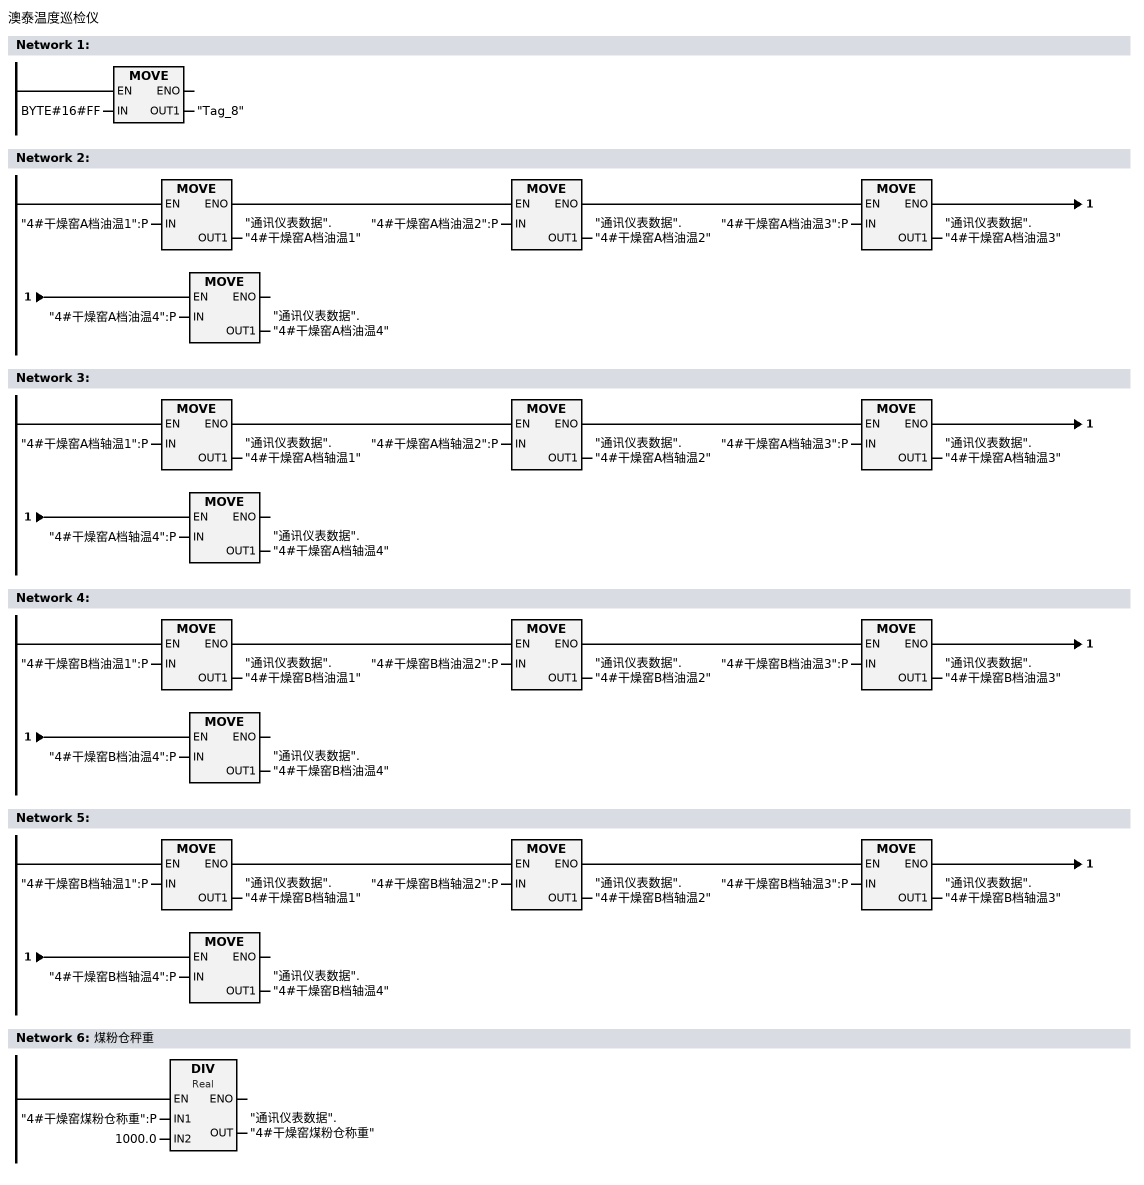
   RUNG wire#powerrail
      { S7_GenerateENO := "TRUE" } Move(in := BYTE#16#FF, out1 => "Tag_8")
   END_RUNG
   // the same network as SCL:
   "Tag_8" := BYTE#16#FF;
END_REGION

REGION Network 2
   RUNG wire#powerrail
      { S7_GenerateENO := "TRUE" } Move(in := "4#干燥窑A档油温1":P, out1 => "通讯仪表数据"."4#干燥窑A档油温1")
      { S7_GenerateENO := "TRUE" } Move(in := "4#干燥窑A档油温2":P, out1 => "通讯仪表数据"."4#干燥窑A档油温2")
      { S7_GenerateENO := "TRUE" } Move(in := "4#干燥窑A档油温3":P, out1 => "通讯仪表数据"."4#干燥窑A档油温3")
      { S7_GenerateENO := "TRUE" } Move(in := "4#干燥窑A档油温4":P, out1 => "通讯仪表数据"."4#干燥窑A档油温4")
   END_RUNG
   // the same network as SCL:
   // ENO of a box is taken as its EN; it also drops when the box reports an error
   "通讯仪表数据"."4#干燥窑A档油温1" := "4#干燥窑A档油温1":P;
   "通讯仪表数据"."4#干燥窑A档油温2" := "4#干燥窑A档油温2":P;
   "通讯仪表数据"."4#干燥窑A档油温3" := "4#干燥窑A档油温3":P;
   "通讯仪表数据"."4#干燥窑A档油温4" := "4#干燥窑A档油温4":P;
END_REGION

REGION Network 3
   RUNG wire#powerrail
      { S7_GenerateENO := "TRUE" } Move(in := "4#干燥窑A档轴温1":P, out1 => "通讯仪表数据"."4#干燥窑A档轴温1")
      { S7_GenerateENO := "TRUE" } Move(in := "4#干燥窑A档轴温2":P, out1 => "通讯仪表数据"."4#干燥窑A档轴温2")
      { S7_GenerateENO := "TRUE" } Move(in := "4#干燥窑A档轴温3":P, out1 => "通讯仪表数据"."4#干燥窑A档轴温3")
      { S7_GenerateENO := "TRUE" } Move(in := "4#干燥窑A档轴温4":P, out1 => "通讯仪表数据"."4#干燥窑A档轴温4")
   END_RUNG
   // the same network as SCL:
   // ENO of a box is taken as its EN; it also drops when the box reports an error
   "通讯仪表数据"."4#干燥窑A档轴温1" := "4#干燥窑A档轴温1":P;
   "通讯仪表数据"."4#干燥窑A档轴温2" := "4#干燥窑A档轴温2":P;
   "通讯仪表数据"."4#干燥窑A档轴温3" := "4#干燥窑A档轴温3":P;
   "通讯仪表数据"."4#干燥窑A档轴温4" := "4#干燥窑A档轴温4":P;
END_REGION

REGION Network 4
   RUNG wire#powerrail
      { S7_GenerateENO := "TRUE" } Move(in := "4#干燥窑B档油温1":P, out1 => "通讯仪表数据"."4#干燥窑B档油温1")
      { S7_GenerateENO := "TRUE" } Move(in := "4#干燥窑B档油温2":P, out1 => "通讯仪表数据"."4#干燥窑B档油温2")
      { S7_GenerateENO := "TRUE" } Move(in := "4#干燥窑B档油温3":P, out1 => "通讯仪表数据"."4#干燥窑B档油温3")
      { S7_GenerateENO := "TRUE" } Move(in := "4#干燥窑B档油温4":P, out1 => "通讯仪表数据"."4#干燥窑B档油温4")
   END_RUNG
   // the same network as SCL:
   // ENO of a box is taken as its EN; it also drops when the box reports an error
   "通讯仪表数据"."4#干燥窑B档油温1" := "4#干燥窑B档油温1":P;
   "通讯仪表数据"."4#干燥窑B档油温2" := "4#干燥窑B档油温2":P;
   "通讯仪表数据"."4#干燥窑B档油温3" := "4#干燥窑B档油温3":P;
   "通讯仪表数据"."4#干燥窑B档油温4" := "4#干燥窑B档油温4":P;
END_REGION

REGION Network 5
   RUNG wire#powerrail
      { S7_GenerateENO := "TRUE" } Move(in := "4#干燥窑B档轴温1":P, out1 => "通讯仪表数据"."4#干燥窑B档轴温1")
      { S7_GenerateENO := "TRUE" } Move(in := "4#干燥窑B档轴温2":P, out1 => "通讯仪表数据"."4#干燥窑B档轴温2")
      { S7_GenerateENO := "TRUE" } Move(in := "4#干燥窑B档轴温3":P, out1 => "通讯仪表数据"."4#干燥窑B档轴温3")
      { S7_GenerateENO := "TRUE" } Move(in := "4#干燥窑B档轴温4":P, out1 => "通讯仪表数据"."4#干燥窑B档轴温4")
   END_RUNG
   // the same network as SCL:
   // ENO of a box is taken as its EN; it also drops when the box reports an error
   "通讯仪表数据"."4#干燥窑B档轴温1" := "4#干燥窑B档轴温1":P;
   "通讯仪表数据"."4#干燥窑B档轴温2" := "4#干燥窑B档轴温2":P;
   "通讯仪表数据"."4#干燥窑B档轴温3" := "4#干燥窑B档轴温3":P;
   "通讯仪表数据"."4#干燥窑B档轴温4" := "4#干燥窑B档轴温4":P;
END_REGION

REGION Network 6: 煤粉仓秤重
   RUNG wire#powerrail
      { S7_Templates := "SrcType := Real" } Div(in1 := "4#干燥窑煤粉仓称重":P, in2 := 1000.0, out => "通讯仪表数据"."4#干燥窑煤粉仓称重")
   END_RUNG
   // the same network as SCL:
   "通讯仪表数据"."4#干燥窑煤粉仓称重" := "4#干燥窑煤粉仓称重":P / 1000.0;
END_REGION
END_FUNCTION

FUNCTION "3#4#干燥窑皮带联锁信号通" : Void   // FC16, LAD
{ S7_Optimized_Access := 'FALSE' }
VERSION : 0.1
BEGIN

REGION Network 1
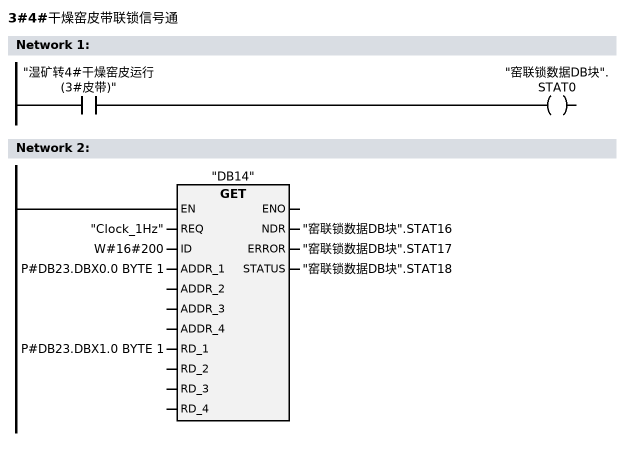
   RUNG wire#powerrail
      Contact( "湿矿转4#干燥窑皮运行  (3#皮带)" )
      Coil( "窑联锁数据DB块".STAT0 )
   END_RUNG
   // the same network as SCL:
   "窑联锁数据DB块".STAT0 := "湿矿转4#干燥窑皮运行  (3#皮带)";
END_REGION

REGION Network 2
   "DB14"(REQ := "Clock_1Hz",   // GET
          ID := W#16#200,
          ADDR_1 := P#DB23.DBX0.0 BYTE 1,
          RD_1 := P#DB23.DBX1.0 BYTE 1,
          NDR => "窑联锁数据DB块".STAT16,
          ERROR => "窑联锁数据DB块".STAT17,
          STATUS => "窑联锁数据DB块".STAT18);
END_REGION
END_FUNCTION

FUNCTION "模拟量转换" : Void   // FC21, LAD
{ S7_Optimized_Access := 'FALSE' }
VERSION : 0.1
BEGIN

REGION Network 1
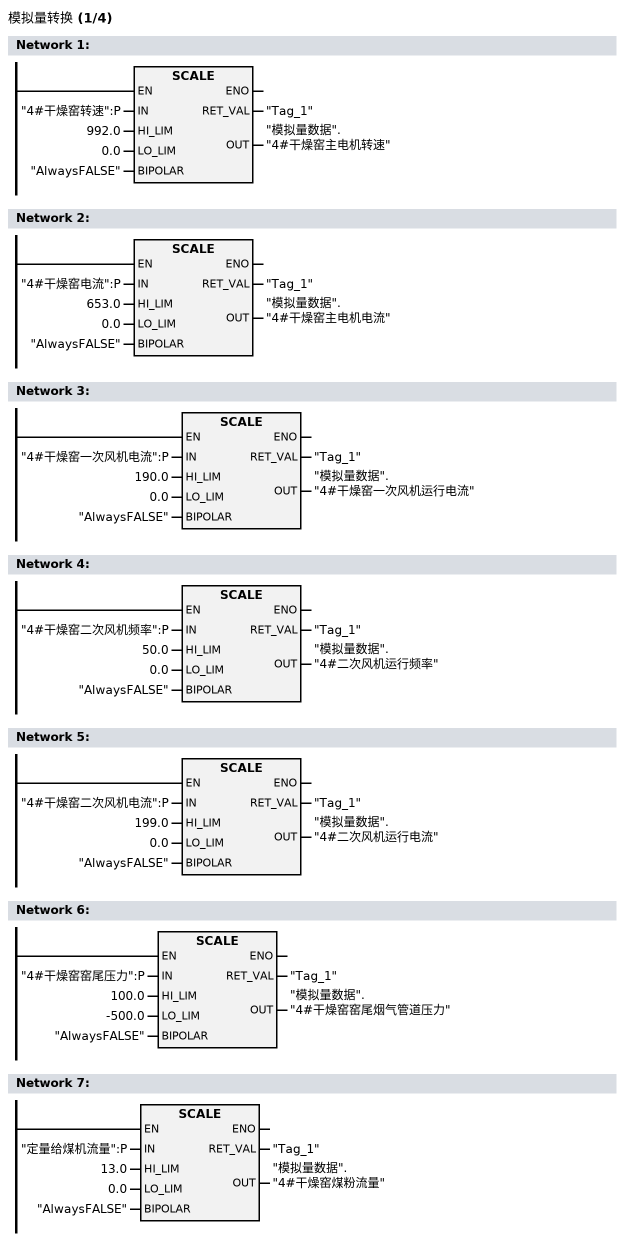
   "Tag_1" := SCALE(IN := "4#干燥窑转速":P,
                    HI_LIM := 992.0,
                    LO_LIM := 0.0,
                    BIPOLAR := "AlwaysFALSE",
                    OUT => "模拟量数据"."4#干燥窑主电机转速");
END_REGION

REGION Network 2
   "Tag_1" := SCALE(IN := "4#干燥窑电流":P,
                    HI_LIM := 653.0,
                    LO_LIM := 0.0,
                    BIPOLAR := "AlwaysFALSE",
                    OUT => "模拟量数据"."4#干燥窑主电机电流");
END_REGION

REGION Network 3
   "Tag_1" := SCALE(IN := "4#干燥窑一次风机电流":P,
                    HI_LIM := 190.0,
                    LO_LIM := 0.0,
                    BIPOLAR := "AlwaysFALSE",
                    OUT => "模拟量数据"."4#干燥窑一次风机运行电流");
END_REGION

REGION Network 4
   "Tag_1" := SCALE(IN := "4#干燥窑二次风机频率":P,
                    HI_LIM := 50.0,
                    LO_LIM := 0.0,
                    BIPOLAR := "AlwaysFALSE",
                    OUT => "模拟量数据"."4#二次风机运行频率");
END_REGION

REGION Network 5
   "Tag_1" := SCALE(IN := "4#干燥窑二次风机电流":P,
                    HI_LIM := 199.0,
                    LO_LIM := 0.0,
                    BIPOLAR := "AlwaysFALSE",
                    OUT => "模拟量数据"."4#二次风机运行电流");
END_REGION

REGION Network 6
   "Tag_1" := SCALE(IN := "4#干燥窑窑尾压力":P,
                    HI_LIM := 100.0,
                    LO_LIM := -500.0,
                    BIPOLAR := "AlwaysFALSE",
                    OUT => "模拟量数据"."4#干燥窑窑尾烟气管道压力");
END_REGION

REGION Network 7
   "Tag_1" := SCALE(IN := "定量给煤机流量":P,
                    HI_LIM := 13.0,
                    LO_LIM := 0.0,
                    BIPOLAR := "AlwaysFALSE",
                    OUT => "模拟量数据"."4#干燥窑煤粉流量");
END_REGION

REGION Network 8
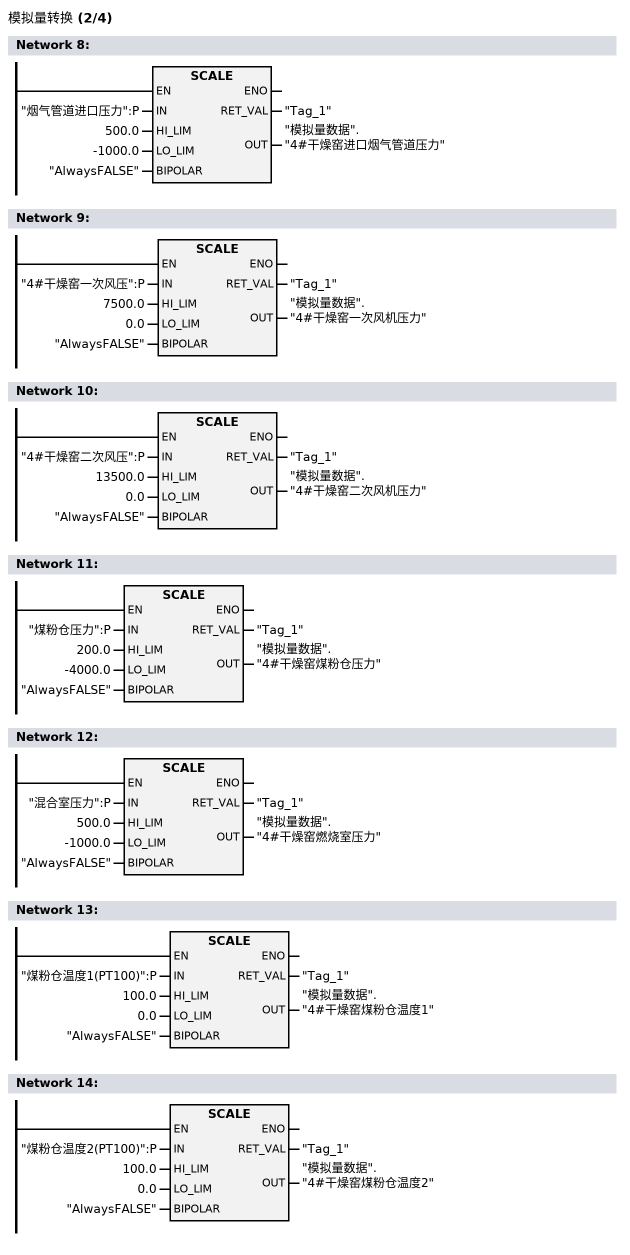
   "Tag_1" := SCALE(IN := "烟气管道进口压力":P,
                    HI_LIM := 500.0,
                    LO_LIM := -1000.0,
                    BIPOLAR := "AlwaysFALSE",
                    OUT => "模拟量数据"."4#干燥窑进口烟气管道压力");
END_REGION

REGION Network 9
   "Tag_1" := SCALE(IN := "4#干燥窑一次风压":P,
                    HI_LIM := 7500.0,
                    LO_LIM := 0.0,
                    BIPOLAR := "AlwaysFALSE",
                    OUT => "模拟量数据"."4#干燥窑一次风机压力");
END_REGION

REGION Network 10
   "Tag_1" := SCALE(IN := "4#干燥窑二次风压":P,
                    HI_LIM := 13500.0,
                    LO_LIM := 0.0,
                    BIPOLAR := "AlwaysFALSE",
                    OUT => "模拟量数据"."4#干燥窑二次风机压力");
END_REGION

REGION Network 11
   "Tag_1" := SCALE(IN := "煤粉仓压力":P,
                    HI_LIM := 200.0,
                    LO_LIM := -4000.0,
                    BIPOLAR := "AlwaysFALSE",
                    OUT => "模拟量数据"."4#干燥窑煤粉仓压力");
END_REGION

REGION Network 12
   "Tag_1" := SCALE(IN := "混合室压力":P,
                    HI_LIM := 500.0,
                    LO_LIM := -1000.0,
                    BIPOLAR := "AlwaysFALSE",
                    OUT => "模拟量数据"."4#干燥窑燃烧室压力");
END_REGION

REGION Network 13
   "Tag_1" := SCALE(IN := "煤粉仓温度1(PT100)":P,
                    HI_LIM := 100.0,
                    LO_LIM := 0.0,
                    BIPOLAR := "AlwaysFALSE",
                    OUT => "模拟量数据"."4#干燥窑煤粉仓温度1");
END_REGION

REGION Network 14
   "Tag_1" := SCALE(IN := "煤粉仓温度2(PT100)":P,
                    HI_LIM := 100.0,
                    LO_LIM := 0.0,
                    BIPOLAR := "AlwaysFALSE",
                    OUT => "模拟量数据"."4#干燥窑煤粉仓温度2");
END_REGION

REGION Network 15
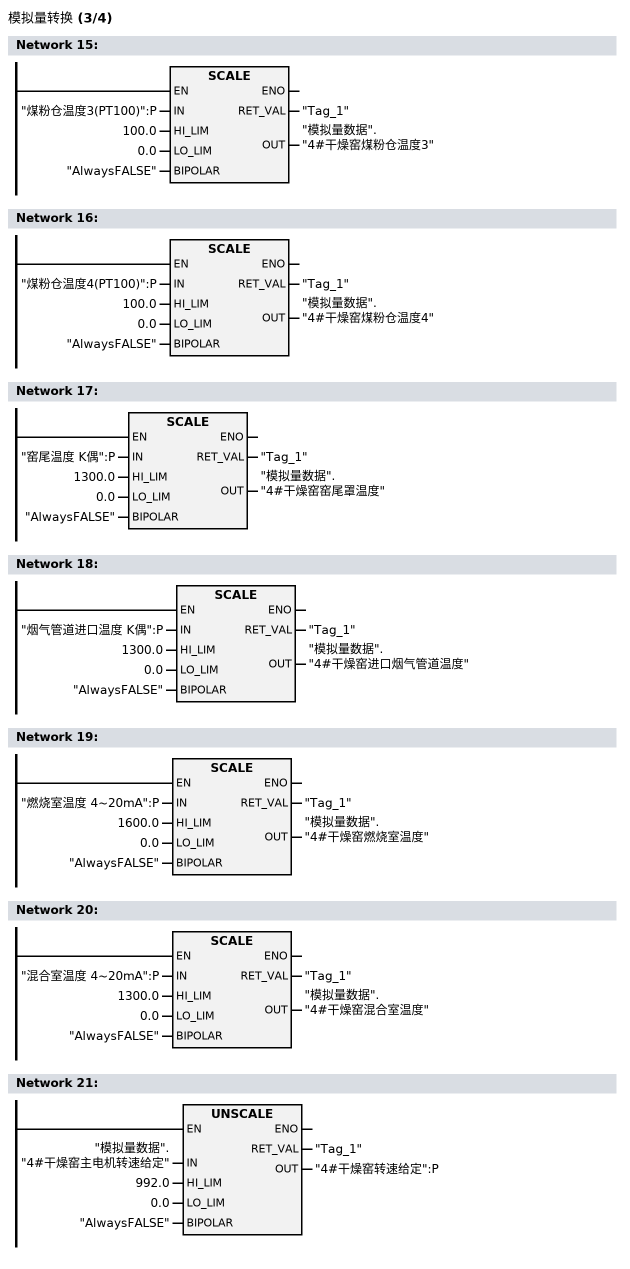
   "Tag_1" := SCALE(IN := "煤粉仓温度3(PT100)":P,
                    HI_LIM := 100.0,
                    LO_LIM := 0.0,
                    BIPOLAR := "AlwaysFALSE",
                    OUT => "模拟量数据"."4#干燥窑煤粉仓温度3");
END_REGION

REGION Network 16
   "Tag_1" := SCALE(IN := "煤粉仓温度4(PT100)":P,
                    HI_LIM := 100.0,
                    LO_LIM := 0.0,
                    BIPOLAR := "AlwaysFALSE",
                    OUT => "模拟量数据"."4#干燥窑煤粉仓温度4");
END_REGION

REGION Network 17
   "Tag_1" := SCALE(IN := "窑尾温度 K偶":P,
                    HI_LIM := 1300.0,
                    LO_LIM := 0.0,
                    BIPOLAR := "AlwaysFALSE",
                    OUT => "模拟量数据"."4#干燥窑窑尾罩温度");
END_REGION

REGION Network 18
   "Tag_1" := SCALE(IN := "烟气管道进口温度 K偶":P,
                    HI_LIM := 1300.0,
                    LO_LIM := 0.0,
                    BIPOLAR := "AlwaysFALSE",
                    OUT => "模拟量数据"."4#干燥窑进口烟气管道温度");
END_REGION

REGION Network 19
   "Tag_1" := SCALE(IN := "燃烧室温度 4~20mA":P,
                    HI_LIM := 1600.0,
                    LO_LIM := 0.0,
                    BIPOLAR := "AlwaysFALSE",
                    OUT => "模拟量数据"."4#干燥窑燃烧室温度");
END_REGION

REGION Network 20
   "Tag_1" := SCALE(IN := "混合室温度 4~20mA":P,
                    HI_LIM := 1300.0,
                    LO_LIM := 0.0,
                    BIPOLAR := "AlwaysFALSE",
                    OUT => "模拟量数据"."4#干燥窑混合室温度");
END_REGION

REGION Network 21
   "Tag_1" := UNSCALE(IN := "模拟量数据"."4#干燥窑主电机转速给定",
                      HI_LIM := 992.0,
                      LO_LIM := 0.0,
                      BIPOLAR := "AlwaysFALSE",
                      OUT => "4#干燥窑转速给定":P);
END_REGION

REGION Network 22
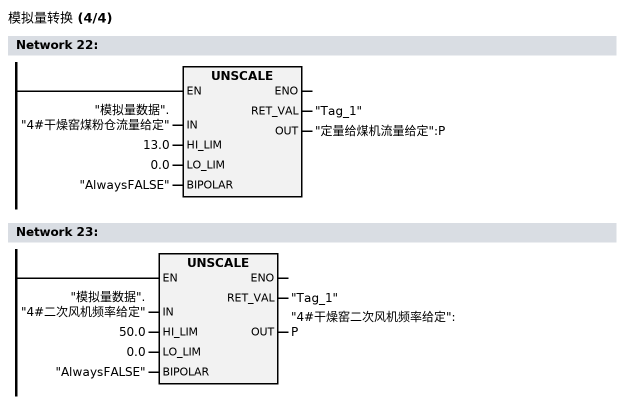
   "Tag_1" := UNSCALE(IN := "模拟量数据"."4#干燥窑煤粉仓流量给定",
                      HI_LIM := 13.0,
                      LO_LIM := 0.0,
                      BIPOLAR := "AlwaysFALSE",
                      OUT => "定量给煤机流量给定":P);
END_REGION

REGION Network 23
   "Tag_1" := UNSCALE(IN := "模拟量数据"."4#二次风机频率给定",
                      HI_LIM := 50.0,
                      LO_LIM := 0.0,
                      BIPOLAR := "AlwaysFALSE",
                      OUT => "4#干燥窑二次风机频率给定":P);
END_REGION
END_FUNCTION

FUNCTION "FC23" : Void   // FC23, LAD
{ S7_Optimized_Access := 'FALSE' }
VERSION : 0.1
   VAR_TEMP   // added for the SCL form of the ladder/FBD networks
      _w1 : Bool;
      _w2 : Bool;
   END_VAR
BEGIN

REGION Network 1
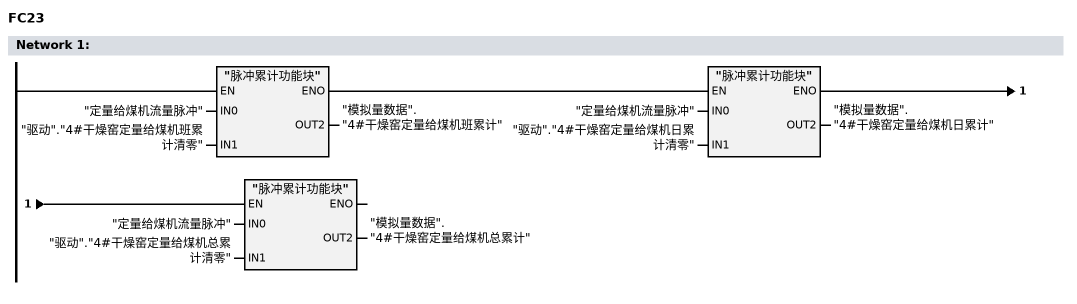
   RUNG wire#powerrail
      "脉冲累计功能块"(IN0 := "定量给煤机流量脉冲", IN1 := "驱动"."4#干燥窑定量给煤机班累计清零", OUT2 => "模拟量数据"."4#干燥窑定量给煤机班累计")
      "脉冲累计功能块"(IN0 := "定量给煤机流量脉冲", IN1 := "驱动"."4#干燥窑定量给煤机日累计清零", OUT2 => "模拟量数据"."4#干燥窑定量给煤机日累计")
      "脉冲累计功能块"(IN0 := "定量给煤机流量脉冲", IN1 := "驱动"."4#干燥窑定量给煤机总累计清零", OUT2 => "模拟量数据"."4#干燥窑定量给煤机总累计")
   END_RUNG
   // the same network as SCL:
   "脉冲累计功能块"(IN0 := "定量给煤机流量脉冲", IN1 := "驱动"."4#干燥窑定量给煤机班累计清零", OUT2 => "模拟量数据"."4#干燥窑定量给煤机班累计", ENO => #_w1);
   "脉冲累计功能块"(EN := #_w1,
             IN0 := "定量给煤机流量脉冲",
             IN1 := "驱动"."4#干燥窑定量给煤机日累计清零",
             OUT2 => "模拟量数据"."4#干燥窑定量给煤机日累计",
             ENO => #_w2);
   IF #_w2 THEN
       "脉冲累计功能块"(IN0 := "定量给煤机流量脉冲", IN1 := "驱动"."4#干燥窑定量给煤机总累计清零", OUT2 => "模拟量数据"."4#干燥窑定量给煤机总累计");
   END_IF;
END_REGION
END_FUNCTION

FUNCTION "FC40_DATA_ALARM" : Void   // FC40, LAD
{ S7_Optimized_Access := 'TRUE' }
VERSION : 0.1
BEGIN

REGION Network 1
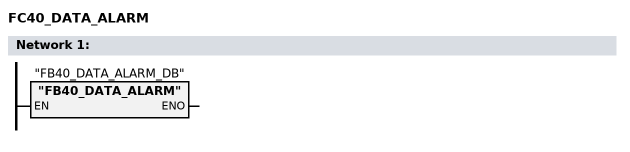
   RUNG wire#powerrail
      "FB40_DATA_ALARM_DB"()
   END_RUNG
   // the same network as SCL:
   "FB40_DATA_ALARM_DB"();   // "FB40_DATA_ALARM"
END_REGION
END_FUNCTION

FUNCTION "脉冲累计功能块" : Void   // FC116, LAD
{ S7_Optimized_Access := 'FALSE' }
VERSION : 0.1
   VAR_INPUT
      IN0 : Bool;
      IN1 : Bool;
   END_VAR
   VAR_OUTPUT
      OUT2 : Real;
   END_VAR
   VAR_TEMP
      TEMP3 : Bool;
      TEMP4 : Real;
      TEMP5 : Real;
      TEMP6 : Real;
   END_VAR
   VAR_TEMP   // added for the SCL form of the ladder/FBD networks
      _w1 : Bool;
   END_VAR
BEGIN

REGION Network 2
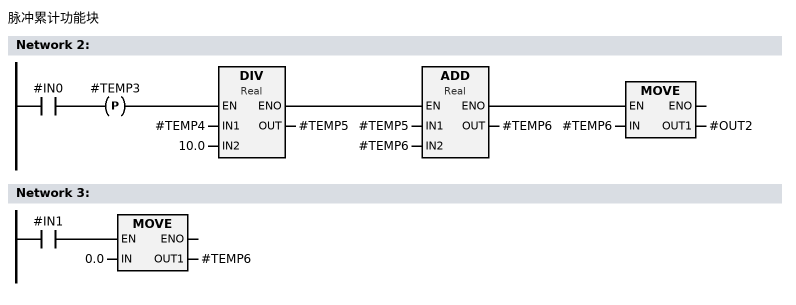
   RUNG wire#powerrail
      Contact( #IN0 )
      P_Trig( #TEMP3 )
      { S7_Templates := "SrcType := Real"; S7_GenerateENO := "TRUE" } Div(in1 := #TEMP4, in2 := 10.0, out => #TEMP5)
      { S7_Templates := "SrcType := Real"; S7_GenerateENO := "TRUE" } Add(in1 := #TEMP5, in2 := #TEMP6, out => #TEMP6)
      { S7_GenerateENO := "TRUE" } Move(in := #TEMP6, out1 => #OUT2)
   END_RUNG
   // the same network as SCL:
   // ENO of a box is taken as its EN; it also drops when the box reports an error
   #_w1 := #IN0 AND NOT #TEMP3;   // rising edge
   #TEMP3 := #IN0;
   IF #_w1 THEN
       #TEMP5 := #TEMP4 / 10.0;
       #TEMP6 := #TEMP5 + #TEMP6;
       #OUT2 := #TEMP6;
   END_IF;
END_REGION

REGION Network 3
   RUNG wire#powerrail
      Contact( #IN1 )
      { S7_GenerateENO := "TRUE" } Move(in := 0.0, out1 => #TEMP6)
   END_RUNG
   // the same network as SCL:
   IF #IN1 THEN #TEMP6 := 0.0; END_IF;
END_REGION

REGION Network 4 (STL)
         SET;
         SAVE;
END_REGION
END_FUNCTION

ORGANIZATION_BLOCK "Main"   // OB1, LAD, ProgramCycle
{ S7_Optimized_Access := 'FALSE' }
VERSION : 0.1
   VAR_TEMP
      TEMP0 : Byte;
      TEMP1 : Byte;
      TEMP2 : Byte;
      TEMP3 : Byte;
      TEMP4 : Byte;
      TEMP5 : Byte;
      TEMP6 : Int;
      TEMP7 : Int;
      TEMP8 : Int;
      TEMP9 : Date_And_Time;
   END_VAR
BEGIN

REGION Network 1
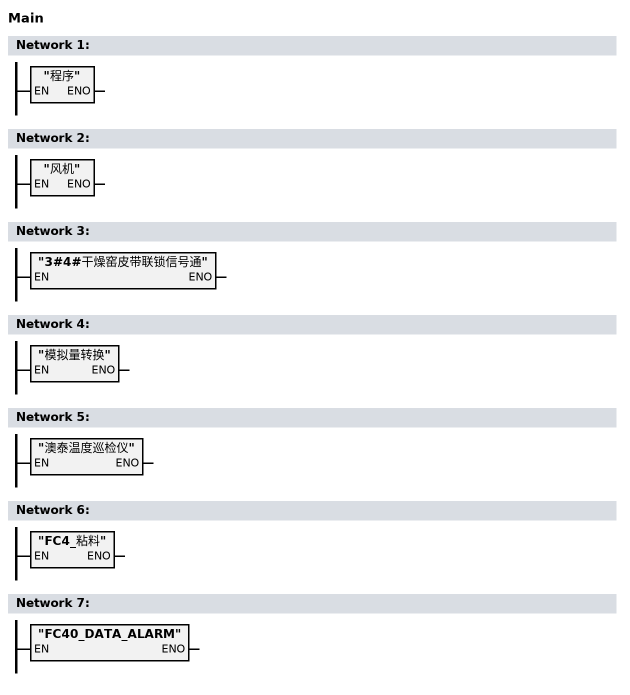
   RUNG wire#powerrail
      "程序"()
   END_RUNG
   // the same network as SCL:
   "程序"();
END_REGION

REGION Network 2
   RUNG wire#powerrail
      "风机"()
   END_RUNG
   // the same network as SCL:
   "风机"();
END_REGION

REGION Network 3
   RUNG wire#powerrail
      "3#4#干燥窑皮带联锁信号通"()
   END_RUNG
   // the same network as SCL:
   "3#4#干燥窑皮带联锁信号通"();
END_REGION

REGION Network 4
   RUNG wire#powerrail
      "模拟量转换"()
   END_RUNG
   // the same network as SCL:
   "模拟量转换"();
END_REGION

REGION Network 5
   RUNG wire#powerrail
      "澳泰温度巡检仪"()
   END_RUNG
   // the same network as SCL:
   "澳泰温度巡检仪"();
END_REGION

REGION Network 6
   RUNG wire#powerrail
      "FC4_粘料"()
   END_RUNG
   // the same network as SCL:
   "FC4_粘料"();
END_REGION

REGION Network 7
   RUNG wire#powerrail
      "FC40_DATA_ALARM"()
   END_RUNG
   // the same network as SCL:
   "FC40_DATA_ALARM"();
END_REGION
END_ORGANIZATION_BLOCK

ORGANIZATION_BLOCK "Cyclic interrupt"   // OB30, LAD, CyclicInterrupt
{ S7_Optimized_Access := 'TRUE' }
VERSION : 0.1
   VAR_INPUT
      Initial_Call : Bool;   // Initial call of this OB
      Event_Count : Int;   // Events discarded
   END_VAR
   VAR_TEMP   // added for the SCL form of the ladder/FBD networks
      _w1 : Bool;
      _w2 : Bool;
   END_VAR
BEGIN

REGION Network 1
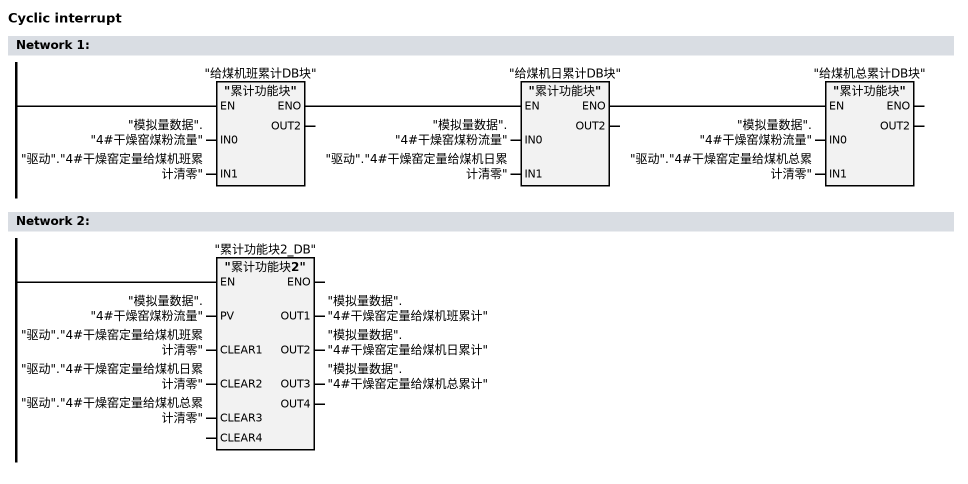
   RUNG wire#powerrail
      "给煤机班累计DB块"(IN0 := "模拟量数据"."4#干燥窑煤粉流量", IN1 := "驱动"."4#干燥窑定量给煤机班累计清零", OUT2 =>)
      "给煤机日累计DB块"(IN0 := "模拟量数据"."4#干燥窑煤粉流量", IN1 := "驱动"."4#干燥窑定量给煤机日累计清零", OUT2 =>)
      "给煤机总累计DB块"(IN0 := "模拟量数据"."4#干燥窑煤粉流量", IN1 := "驱动"."4#干燥窑定量给煤机总累计清零", OUT2 =>)
   END_RUNG
   // the same network as SCL:
   "给煤机班累计DB块"(IN0 := "模拟量数据"."4#干燥窑煤粉流量", IN1 := "驱动"."4#干燥窑定量给煤机班累计清零", ENO => #_w1);   // "累计功能块"
   "给煤机日累计DB块"(EN := #_w1, IN0 := "模拟量数据"."4#干燥窑煤粉流量", IN1 := "驱动"."4#干燥窑定量给煤机日累计清零", ENO => #_w2);   // "累计功能块"
   IF #_w2 THEN
       "给煤机总累计DB块"(IN0 := "模拟量数据"."4#干燥窑煤粉流量", IN1 := "驱动"."4#干燥窑定量给煤机总累计清零");   // "累计功能块"
   END_IF;
END_REGION

REGION Network 2
   RUNG wire#powerrail
      "累计功能块2_DB"(PV := "模拟量数据"."4#干燥窑煤粉流量", CLEAR1 := "驱动"."4#干燥窑定量给煤机班累计清零", CLEAR2 := "驱动"."4#干燥窑定量给煤机日累计清零", CLEAR3 := "驱动"."4#干燥窑定量给煤机总累计清零", CLEAR4 :=, OUT1 => "模拟量数据"."4#干燥窑定量给煤机班累计", OUT2 => "模拟量数据"."4#干燥窑定量给煤机日累计", OUT3 => "模拟量数据"."4#干燥窑定量给煤机总累计", OUT4 =>)
   END_RUNG
   // the same network as SCL:
   "累计功能块2_DB"(PV := "模拟量数据"."4#干燥窑煤粉流量",   // "累计功能块2"
               CLEAR1 := "驱动"."4#干燥窑定量给煤机班累计清零",
               CLEAR2 := "驱动"."4#干燥窑定量给煤机日累计清零",
               CLEAR3 := "驱动"."4#干燥窑定量给煤机总累计清零",
               OUT1 => "模拟量数据"."4#干燥窑定量给煤机班累计",
               OUT2 => "模拟量数据"."4#干燥窑定量给煤机日累计",
               OUT3 => "模拟量数据"."4#干燥窑定量给煤机总累计");
END_REGION
END_ORGANIZATION_BLOCK

// ===== PLC "4#HZY"  CPU 1511-1 PN =====

VAR_GLOBAL   // PLC tag table "默认变量表"
   "转子秤运行" AT %I8.1 : Bool;
   "转子秤流量脉冲" AT %I8.3 : Bool;
   "转子秤流量反馈" AT %IW302 : Int;
   "转子秤故障" AT %I8.2 : Bool;
   "转子秤中控" AT %I8.0 : Bool;
   "窑尾温度K偶" AT %IW280 : Int;
   "窑尾压力" AT %IW264 : Int;
   "窑头温度" AT %IW322 : Int;
   "窑体行程下限" AT %I5.2 : Bool;
   "窑体行程下下限" AT %I5.3 : Bool;
   "窑体行程上限" AT %I5.0 : Bool;
   "窑体行程上上限" AT %I5.1 : Bool;
   "窑体温度6" AT %IW334 : Int;
   "窑体温度5" AT %IW332 : Int;
   "窑体温度4" AT %IW330 : Int;
   "窑体温度3" AT %IW328 : Int;
   "窑体温度2" AT %IW326 : Int;
   "窑体温度1" AT %IW324 : Int;
   "煤粉仓负压" AT %IW300 : Int;
   "回转窑助燃罗茨风机电流" AT %IW320 : Int;
   "回转窑助燃罗茨风机频率" AT %IW318 : Int;
   "煤粉仓温度4" AT %IW316 : Int;
   "煤粉仓温度3" AT %IW314 : Int;
   "煤粉仓温度2" AT %IW312 : Int;
   "煤粉仓温度1" AT %IW310 : Int;
   "煤粉仓收尘风机运行" AT %I8.5 : Bool;
   "煤粉仓收尘风机故障" AT %I8.6 : Bool;
   "煤粉仓收尘风机中控" AT %I8.4 : Bool;
   "烟道闸阀标尺" AT %IW270 : Int;
   "板式给料机流量" AT %IW350 : Int;
   "挡轮重故障" AT %I4.4 : Bool;
   "挡轮轻故障" AT %I4.5 : Bool;
   "干矿进料皮带运行" AT %I6.4 : Bool;
   "干矿进料皮带故障" AT %I6.5 : Bool;
   "干矿进料皮带中控" AT %I6.3 : Bool;
   "干矿提升皮带运行" AT %I6.1 : Bool;
   "干矿提升皮带故障" AT %I6.2 : Bool;
   "干矿提升皮带中控" AT %I6.0 : Bool;
   "尾排风机高压远程" AT %I7.0 : Bool;
   "尾排风机高压合闸" AT %I7.1 : Bool;
   "尾排风机高压分闸" AT %I7.2 : Bool;
   "尾排风机频率反馈" AT %IW268 : Int;
   "尾排风机电流反馈" AT %IW266 : Int;
   "尾排风机变频远程" AT %I7.4 : Bool;
   "尾排风机变频运行" AT %I7.5 : Bool;
   "尾排风机变频故障" AT %I7.6 : Bool;
   "尾排风机变频待机" AT %I7.7 : Bool;
   "回转窑窑头护板风机运行" AT %I11.1 : Bool;
   "回转窑窑头护板风机故障" AT %I11.2 : Bool;
   "回转窑窑头护板风机中控" AT %I11.0 : Bool;
   "回转窑窑头压力" AT %IW304 : Int;
   "回转窑备用风机频率" AT %IW296 : Int;
   "回转窑备用风机电流" AT %IW298 : Int;
   "4#回转窑富氧快切阀关到位" AT %I10.4 : Bool;
   "回转窑备用二次风机故障" AT %I10.5 : Bool;
   "4#回转窑富氧快切阀开到位" AT %I10.3 : Bool;
   "回转窑备用一次风机运行" AT %I10.1 : Bool;
   "回转窑备用一次风机故障" AT %I10.2 : Bool;
   "回转窑备用一次风机中控" AT %I10.0 : Bool;
   "回转窑二次风机频率" AT %IW292 : Int;
   "回转窑二次风机运行" AT %I9.4 : Bool;
   "回转窑二次风机电流" AT %IW294 : Int;
   "回转窑二次风机故障" AT %I9.5 : Bool;
   "回转窑二次风机中控" AT %I9.3 : Bool;
   "回转窑一次风机频率" AT %IW288 : Int;
   "回转窑一次风机运行" AT %I9.1 : Bool;
   "回转窑一次风机电流" AT %IW290 : Int;
   "回转窑一次风机故障" AT %I9.2 : Bool;
   "回转窑一次风机中控" AT %I9.0 : Bool;
   "从机转速" AT %IW260 : Int;
   "从机稀油重故障" AT %I3.6 : Bool;
   "从机稀油轻故障" AT %I3.7 : Bool;
   "从机稀油油差下限" AT %I3.3 : Bool;
   "从机稀油油位下限" AT %I3.5 : Bool;
   "从机稀油油位上限" AT %I3.4 : Bool;
   "从机稀油允许主机启动" AT %I5.5 : Bool;
   "从机稀油中控" AT %I3.0 : Bool;
   "从机稀油2#泵运行" AT %I3.2 : Bool;
   "从机稀油1#泵运行" AT %I3.1 : Bool;
   "从机电流" AT %IW262 : Int;
   "二次风压力" AT %IW308 : Int;
   "主机转速" AT %IW256 : Int;
   "主机稀油重故障" AT %I2.6 : Bool;
   "主机稀油轻故障" AT %I2.7 : Bool;
   "主机稀油油差下限" AT %I2.3 : Bool;
   "主机稀油油位下限" AT %I2.5 : Bool;
   "主机稀油油位上限" AT %I2.4 : Bool;
   "主机稀油允许主机启动" AT %I5.4 : Bool;
   "主机稀油中控" AT %I2.0 : Bool;
   "主机稀油2#泵运行" AT %I2.2 : Bool;
   "主机稀油1#泵运行" AT %I2.1 : Bool;
   "主机电流" AT %IW258 : Int;
   "一次风压力" AT %IW306 : Int;
   "从电机后轴温度" AT %IW286 : Int;
   "从电机前轴温度" AT %IW284 : Int;
   "从电机定子温度" AT %IW282 : Int;
   "PIW278" AT %IW278 : Int;
   "主电机后轴温度" AT %IW276 : Int;
   "主电机前轴温度" AT %IW274 : Int;
   "主电机定子温度" AT %IW272 : Int;
   "I9_7" AT %I9.7 : Bool;
   "I9_6" AT %I9.6 : Bool;
   "I8_7" AT %I8.7 : Bool;
   "I7_3" AT %I7.3 : Bool;
   "I6_7" AT %I6.7 : Bool;
   "I6_6" AT %I6.6 : Bool;
   "I5_7" AT %I5.7 : Bool;
   "I5_6" AT %I5.6 : Bool;
   "I4_7" AT %I4.7 : Bool;
   "I4_6" AT %I4.6 : Bool;
   "I17_7" AT %I17.7 : Bool;
   "I17_6" AT %I17.6 : Bool;
   "I17_5" AT %I17.5 : Bool;
   "I17_4" AT %I17.4 : Bool;
   "I17_3" AT %I17.3 : Bool;
   "I17_2" AT %I17.2 : Bool;
   "I17_1" AT %I17.1 : Bool;
   "I17_0" AT %I17.0 : Bool;
   "I16_7" AT %I16.7 : Bool;
   "I16_6" AT %I16.6 : Bool;
   "I16_5" AT %I16.5 : Bool;
   "I16_4" AT %I16.4 : Bool;
   "I15_7" AT %I15.7 : Bool;
   "I15_6" AT %I15.6 : Bool;
   "I15_5" AT %I15.5 : Bool;
   "I15_4" AT %I15.4 : Bool;
   "I11_7" AT %I11.7 : Bool;
   "24# 煤粉仓消防阀关到位" AT %I11.6 : Bool;
   "回转窑助燃罗茨风机运行" AT %I11.5 : Bool;
   "回转窑助燃罗茨风机故障" AT %I11.4 : Bool;
   "回转窑助燃罗茨风机中控" AT %I11.3 : Bool;
   "24# 煤粉仓消防阀开到位" AT %I10.7 : Bool;
   "24# 煤粉仓消防阀自动位" AT %I10.6 : Bool;
   "I1_7" AT %I1.7 : Bool;
   "I1_6" AT %I1.6 : Bool;
   "I1_5" AT %I1.5 : Bool;
   "I1_4" AT %I1.4 : Bool;
   "I1_3" AT %I1.3 : Bool;
   "4#回转窑急停" AT %I1.2 : Bool;
   "4#窑提升皮带打滑检测" AT %I1.1 : Bool;
   "7#配料皮带运行" AT %I15.1 : Bool;
   "7#配料皮带流量脉冲" AT %I15.3 : Bool;
   "7#配料皮带故障" AT %I15.2 : Bool;
   "7#配料皮带备妥" AT %I15.0 : Bool;
   "7#配料流量" AT %IW348 : Int;
   "6#配料皮带运行" AT %I14.5 : Bool;
   "6#配料皮带流量脉冲" AT %I14.7 : Bool;
   "6#配料皮带故障" AT %I14.6 : Bool;
   "6#配料皮带备妥" AT %I14.4 : Bool;
   "6#配料流量" AT %IW346 : Int;
   "5#配料皮带运行" AT %I14.1 : Bool;
   "5#配料皮带流量脉冲" AT %I14.3 : Bool;
   "5#配料皮带故障" AT %I14.2 : Bool;
   "5#配料皮带备妥" AT %I14.0 : Bool;
   "5#配料流量" AT %IW344 : Int;
   "4#配料皮带运行" AT %I13.5 : Bool;
   "4#配料皮带流量脉冲" AT %I13.7 : Bool;
   "4#配料皮带故障" AT %I13.6 : Bool;
   "4#配料皮带备妥" AT %I13.4 : Bool;
   "4#配料流量" AT %IW342 : Int;
   "3#配料皮带运行" AT %I13.1 : Bool;
   "3#配料皮带流量脉冲" AT %I13.3 : Bool;
   "3#配料皮带故障" AT %I13.2 : Bool;
   "3#配料皮带备妥" AT %I13.0 : Bool;
   "3#配料流量" AT %IW340 : Int;
   "2#配料皮带运行" AT %I12.5 : Bool;
   "2#配料皮带流量脉冲" AT %I12.7 : Bool;
   "2#配料皮带故障" AT %I12.6 : Bool;
   "2#配料皮带备妥" AT %I12.4 : Bool;
   "2#配料流量" AT %IW338 : Int;
   "4#回转窑煤粉仓称重" AT %ID600 : DWord;
   "4#回转窑启动备妥" AT %I0.0 : Bool;
   "4#回转窑从机运行" AT %I0.6 : Bool;
   "4#回转窑从机故障" AT %I0.7 : Bool;
   "4#回转窑从机备妥" AT %I0.5 : Bool;
   "4#回转窑从机合闸" AT %I1.0 : Bool;
   "4#回转窑主机运行" AT %I0.2 : Bool;
   "4#回转窑主机故障" AT %I0.3 : Bool;
   "4#回转窑主机备妥" AT %I0.1 : Bool;
   "4#回转窑主机合闸" AT %I0.4 : Bool;
   "4#回转窑中间仓称重" AT %ID608 : DWord;
   "1#配料皮带运行" AT %I12.1 : Bool;
   "1#配料皮带流量脉冲" AT %I12.3 : Bool;
   "1#配料皮带故障" AT %I12.2 : Bool;
   "1#配料皮带备妥" AT %I12.0 : Bool;
   "1#配料流量" AT %IW336 : Int;
   "1#板式给料机运行" AT %I16.1 : Bool;
   "1#板式给料机流量脉冲" AT %I16.3 : Bool;
   "1#板式给料机故障" AT %I16.2 : Bool;
   "1#板式给料机备妥" AT %I16.0 : Bool;
   "1#挡轮溢流阀运行" AT %I4.3 : Bool;
   "1#挡轮备妥" AT %I4.0 : Bool;
   "1#挡轮2#泵运行" AT %I4.2 : Bool;
   "1#挡轮1#泵运行" AT %I4.1 : Bool;
   "4#回转窑支撑挡轮轴温度D4" AT %ID552 : DWord;
   "4#回转窑支撑挡轮轴温度D3" AT %ID544 : DWord;
   "4#回转窑支撑挡轮轴温度D2" AT %ID536 : DWord;
   "4#回转窑支撑挡轮轴温度D1" AT %ID528 : DWord;
   "4#回转窑支撑挡轮轴温度C4" AT %ID520 : DWord;
   "4#回转窑支撑挡轮轴温度C3" AT %ID512 : DWord;
   "4#回转窑支撑挡轮轴温度C2" AT %ID504 : DWord;
   "4#回转窑支撑挡轮轴温度C1" AT %ID496 : DWord;
   "4#回转窑支撑挡轮轴温度B4" AT %ID456 : DWord;
   "4#回转窑支撑挡轮轴温度B3" AT %ID448 : DWord;
   "4#回转窑支撑挡轮轴温度B2" AT %ID440 : DWord;
   "4#回转窑支撑挡轮轴温度B1" AT %ID432 : DWord;
   "4#回转窑支撑挡轮轴温度A4" AT %ID424 : DWord;
   "4#回转窑支撑挡轮轴温度A3" AT %ID416 : DWord;
   "4#回转窑支撑挡轮轴温度A2" AT %ID408 : DWord;
   "4#回转窑支撑挡轮轴温度A1" AT %ID400 : DWord;
   "4#回转窑支撑挡轮温度D4" AT %ID556 : DWord;
   "4#回转窑支撑挡轮温度D3" AT %ID548 : DWord;
   "4#回转窑支撑挡轮温度D2" AT %ID540 : DWord;
   "4#回转窑支撑挡轮温度D1" AT %ID532 : DWord;
   "4#回转窑支撑挡轮温度C4" AT %ID524 : DWord;
   "4#回转窑支撑挡轮温度C3" AT %ID516 : DWord;
   "4#回转窑支撑挡轮温度C2" AT %ID508 : DWord;
   "4#回转窑支撑挡轮温度C1" AT %ID500 : DWord;
   "4#回转窑支撑挡轮温度B4" AT %ID460 : DWord;
   "4#回转窑支撑挡轮温度B3" AT %ID452 : DWord;
   "4#回转窑支撑挡轮温度B2" AT %ID444 : DWord;
   "4#回转窑支撑挡轮温度B1" AT %ID436 : DWord;
   "4#回转窑支撑挡轮温度A4" AT %ID428 : DWord;
   "4#回转窑支撑挡轮温度A3" AT %ID420 : DWord;
   "4#回转窑支撑挡轮温度A2" AT %ID412 : DWord;
   "4#回转窑支撑挡轮温度A1" AT %ID404 : DWord;
   "转子秤连锁停止" AT %Q5.0 : Bool;
   "转子秤启动" AT %Q4.0 : Bool;
   "给煤机流量给定" AT %QW272 : Int;
   "煤粉仓收尘风机启动" AT %Q4.1 : Bool;
   "板式给料机流量给定" AT %QW302 : Int;
   "板式给料机启动" AT %Q7.0 : Bool;
   "挡轮启动" AT %Q0.4 : Bool;
   "挡轮停止" AT %Q0.7 : Bool;
   "干矿进料皮带启动" AT %Q1.2 : Bool;
   "干矿提升皮带启动" AT %Q1.0 : Bool;
   "尾排风机高压柜变频启动" AT %Q1.5 : Bool;
   "尾排风机高压柜变频停止" AT %Q1.6 : Bool;
   "尾排风机高压合闸驱动" AT %Q1.3 : Bool;
   "尾排风机高压分闸驱动" AT %Q1.4 : Bool;
   "尾排风机频率给定" AT %QW258 : Int;
   "回转窑窑头护板风机启动" AT %Q4.6 : Bool;
   "回转窑备用风机频率给定" AT %QW284 : Int;
   "回转窑备用二次风机启动" AT %Q4.5 : Bool;
   "回转窑备用一次风机启动" AT %Q4.4 : Bool;
   "回转窑合闸" AT %Q0.0 : Bool;
   "回转窑二次风机频率给定" AT %QW282 : Int;
   "回转窑二次风机启动" AT %Q4.3 : Bool;
   "回转窑主机转速给定" AT %QW256 : Int;
   "回转窑主机启动" AT %Q0.1 : Bool;
   "回转窑一次风机频率给定" AT %QW280 : Int;
   "回转窑一次风机启动" AT %Q4.2 : Bool;
   "从机稀油启动" AT %Q0.3 : Bool;
   "从机稀油停止" AT %Q0.6 : Bool;
   "主机稀油启动" AT %Q0.2 : Bool;
   "主机稀油停止" AT %Q0.5 : Bool;
   "Tag_26" AT %QB8 : Byte;
   "3料仓粘仓信号输出" AT %Q7.7 : Bool;
   "2料仓粘仓信号输出" AT %Q7.6 : Bool;
   "1料仓粘仓信号输出" AT %Q7.5 : Bool;
   "7#料仓粘仓信号输出" AT %Q7.4 : Bool;
   "6#料仓粘仓信号输出" AT %Q7.3 : Bool;
   "5#料仓粘仓信号输出" AT %Q7.2 : Bool;
   "4#料仓粘仓信号输出" AT %Q7.1 : Bool;
   "Q6_7" AT %Q6.7 : Bool;
   "4#回转窑富氧快切阀驱动" AT %Q5.7 : Bool;
   "Q5_6" AT %Q5.6 : Bool;
   "Q5_5" AT %Q5.5 : Bool;
   "Q5_4" AT %Q5.4 : Bool;
   "Q5_3" AT %Q5.3 : Bool;
   "24# 煤粉仓消防阀驱动" AT %Q5.2 : Bool;